       IF #Clr AND NOT #edge THEN
           IF #Q0 THEN #Q0 := FALSE;
           ELSIF #Q1 THEN #Q1 := FALSE;
           ELSIF #Q2 THEN #Q2 := FALSE;
           ELSIF #Q3 THEN #Q3 := FALSE;
           ELSIF #Q4 THEN #Q4 := FALSE;
           ELSIF #Q5 THEN #Q5 := FALSE;
           ELSIF #Q6 THEN #Q6 := FALSE;
           ELSE #Q7 := FALSE;
           END_IF;
       END_IF;
       #edge := #Clr;
   END_IF;


   (* revision history
   hm  25.12.2007  rev 1.0
       original version

   hm  30. oct. 2008   rev 1.1
       optimized performance

   hm  14. mar. 2009   rev 1.2
       removed double assignments

   *)
END_FUNCTION_BLOCK

// ===== PLC "Logic Others"  Unspecific CPU S7 300 =====

FUNCTION_BLOCK "CRC_GEN"   // FB72, SCL
TITLE = CRC_GEN
{ S7_Optimized_Access := 'FALSE' }
AUTHOR : hugo
FAMILY : LOGIC
NAME : CRCGEN
VERSION : 2.0
// CRC_GEN generates a CRC checksum from a block of data and returns  the checksum in a DWORD to be connected to the data for transmission.
// the CRC Polynom is specified with the config variable PN and the length of the Polynom is specified by PL
// A Polynom x4 + X + 1 is represented by 0011 with length 4, the highest order bit is not specified at all..
// The input data is an array of byte of any size, the function is called by CRC_GEN(ADR(array),SIZEOF(array), ....).
// 
// uses: REVERSE (FC310)
//       REFLECT (FC426)
   VAR_INPUT
      PT : Pointer;
      _PT AT PT : Struct
         DBNr : Word;
         Adr : DWord;
      END_STRUCT;
      SIZE : Int;
      PL : Int;
      PN : DWord;
      INIT : DWord;
      REV_IN : Bool;
      REV_OUT : Bool;
      XOR_OUT : DWord;
   END_VAR
   VAR_OUTPUT
      CRC_GEN : DWord;
      _CRC_GEN AT CRC_GEN : Array[0..31] of Bool;
   END_VAR
   VAR_TEMP
      pos : Int;
      shift : Int;
      dx : Byte;
      _dx AT dx : Array[0..7] of Bool;
      bits : Int;
      rTEST_DB : Int;
      Adr : Int;
      DB_LENGTH : Word;
      WRITE_PROT : Bool;
   END_VAR
BEGIN


   (* Datenbaustein Testen *)
   #rTEST_DB := TEST_DB(DB_NUMBER := #_PT.DBNr // IN: WORD
                    ,DB_LENGTH => #DB_LENGTH // OUT: WORD
                    ,WRITE_PROT => #WRITE_PROT // OUT: BOOL
                    ); // INT
   (* Ende wenn Test-DB <> 0 = Fehler *)
   IF #rTEST_DB <> 0 THEN RETURN; END_IF;
   (* Ende wenn DB zu klein *) 
   IF WORD_TO_INT(#DB_LENGTH)/1 < #SIZE THEN RETURN; END_IF;

   #Adr := DWORD_TO_INT(SHR(IN:=SHL(IN:=#_PT.Adr,N:=8),N:=11));

   (* align polygon *)
   #shift := 32 - #PL;
   #PN := SHL(IN:=#PN,N:=#shift);

   (* load first 4 bytes into register minimum message size is 4 bytes
     for smaller messages fill with 0#s at the beginning*)
   FOR #pos := 0 TO 3 DO
     IF #REV_IN THEN #CRC_GEN := SHL(IN:=#CRC_GEN,N:=8) OR "REVERSE"(WORD_TO_BLOCK_DB(#_PT.DBNr).DB(#Adr+#pos)); ELSE #CRC_GEN := SHL(IN:=#CRC_GEN,N:=8) OR WORD_TO_BLOCK_DB(#_PT.DBNr).DB(#Adr+#pos); END_IF;
   END_FOR;
   #pos := 4;

   (* xor with init value *)
   #CRC_GEN := #CRC_GEN XOR SHL(IN:=#INIT,N:=#shift);

   (* calculate CRC for each byte *)
   WHILE #pos < #SIZE DO
     IF #REV_IN THEN #dx := "REVERSE"(WORD_TO_BLOCK_DB(#_PT.DBNr).DB(#Adr+#pos)); ELSE #dx := WORD_TO_BLOCK_DB(#_PT.DBNr).DB(#Adr+#pos); END_IF;
     #pos := #pos + 1;
     (* crc calculation for one byte *)
     FOR #bits := 0 TO 7 DO
       IF #_CRC_GEN[7] THEN
         #CRC_GEN := (SHL(IN:=#CRC_GEN,N:=1) OR BOOL_TO_DWORD(#_dx[7])) XOR #PN;
       ELSE
         #CRC_GEN := SHL(IN:=#CRC_GEN,N:=1) OR BOOL_TO_DWORD(#_dx[7]);
       END_IF;
       #dx := SHL(IN:=#dx,N:=1);
     END_FOR;
   END_WHILE;

   (* all bytes are processed, need to finish the registers 32 bits *)
   FOR #bits := 0 TO 31 DO
     IF #_CRC_GEN[7] THEN
       #CRC_GEN := (SHL(IN:=#CRC_GEN,N:=1) OR BOOL_TO_DWORD(#_dx[7])) XOR #PN;
     ELSE
       #CRC_GEN := SHL(IN:=#CRC_GEN,N:=1) OR BOOL_TO_DWORD(#_dx[7]);
     END_IF;
   END_FOR;

   (* final XOR *)
   #CRC_GEN := SHR(IN:=#CRC_GEN,N:=#shift) XOR #XOR_OUT;

   (* reverse the crc_out put if necessary *)
   IF #REV_OUT THEN #CRC_GEN := "REFLECT"(D:=#CRC_GEN,L:=#PL); END_IF;


   (* typical crc polynoms

   CRC-4-ITU       x4 + x + 1          (ITU G.704, p. 12)  0x3 or 0xC (0x9)
   CRC-5-ITU       x5 + x4 + x2 + 1      (ITU G.704, p. 9)   0x15 or 0x15 (0x0B) Bluetooth
   CRC-5-USB       x5 + x2 + 1         (use: USB token packets)  0x05 or 0x14 (0x9)
   CRC-6-ITU       x6 + x + 1          (ITU G.704, p. 3)   0x03 or 0x30 (0x21)
   CRC-7         x7 + x3 + 1         (use: telecom systems, MMC)   0x09 or 0x48 (0x11)
   CRC-8-ATM       x8 + x2 + x + 1         (use: ATM HEC)  0x07 or 0xE0 (0xC1)
   CRC-8-CCITT     x8 + x7 + x3 + x2 + 1     (use: 1-Wire bus)   0x8D or 0xB1 (0x63)
   CRC-8-Dallas/Maxim  x8 + x5 + x4 + 1      (use: 1-Wire bus)   0x31 or 0x8C (0x19)
   CRC-8         x8 + x7 + x6 + x4 + x2 + 1  0xD5 or 0xAB (0x57)
   CRC-8-SAE J1850   x8 + x4 + x3 + x2 + 1     0x1D or 0xB8
   CRC-10        x10 + x9 + x5 + x4 + x + 1  0x233 or 0x331 (0x263)
   CRC-12        x12 + x11 + x3 + x2 + x + 1 (use: telecom systems)   0x80F or 0xF01 (0xE03)
   CRC-15-CAN      x15 + x14 + x10 + x8 + x7 + x4 + x3 + 1   0x4599 or 0x4CD1 (0x19A3)
   CRC-16-Fletcher   Not a CRC; see Fletcher's checksum  Used in Adler-32 A & B CRCs
   CRC-16-CCITT  x16 + x12 + x5 + 1 (XMODEM,X.25, V.41, Bluetooth, PPP, IrDA; known as "CRC-CCITT")  0x1021 or 0x8408 (0x0811)
   CRC-16-IBM  x16 + x15 + x2 + 1 (USB, many others; also known as "CRC-16")   0x8005 or 0xA001 (0x4003)
   CRC-24-Radix-64   x24 + x23 + x18 + x17 + x14 + x11 + x10 + x7 + x6 + x5 + x4 + x3 + x + 1  0x864CFB or 0xDF3261 (0xBE64C3)
   CRC-32-Adler  Not a CRC; see Adler-32   See Adler-32
   CRC-32-MPEG2  x32 + x26 + x23 + x22 + x16 + x12 + x11 + x10 + x8 + x7 + x5 + x4 + x2 + x + 1  0x04C11DB7 or 0xEDB88320 (0xDB710641) Also used in IEEE 802.3
   CRC-32-IEEE 802.3   x32 + x26 + x23 + x22 + x16 + x12 + x11 + x10 + x8 + x7 + x5 + x4 + x2 + x + 1 (V.42)   0x04C11DB7 or 0xEDB88320 (0xDB710641)
   CRC-32C (Castagnoli)  x32 + x28 + x27 + x26 + x25 + x23 + x22 + x20 + x19 + x18 + x14 + x13 + x11 + x10 + x9 + x8 + x6 + 1  0x1EDC6F41 or 0x82F63B78 (0x05EC76F1)
   CRC-64-ISO  x64 + x4 + x3 + x + 1 (use: ISO 3309)   0x000000000000001B or 0xD800000000000000 (0xB000000000000001)
   CRC-64-ECMA-182   x64 + x62 + x57 + x55 + x54 + x53 + x52 + x47 + x46 + x45 + x40 + x39 + x38 + x37 + x35 + x33 + x32 + x31 + x29 + x27 + x24 + x23 + x22 + x21 + x19 + x17 + x13 + x12 + x10 + x9 + x7 + x4 + x + 1
   (as described in ECMA-182 p.63)   0x42F0E1EBA9EA3693 or 0xC96C5795D7870F42 (0x92D8AF2BAF0E1E85)
   *)



   (* revision history

   hm  9.6.2007    rev 1.0   
     original version 

   hm  11.9.2007   rev 1.1
     deleted unused variable i

   hm  9. oct 2007   rev 1.2
     added init code for crc and xor_out
     added refelct in and reflect_out (rev_in und Rev_out)

   hm  2. jan 2008 rev 1.3
     small changes for performance improvements

   hm  16. mar. 2008 rev 1.4
     changed type of input size to uint

   hm  10. mar. 2009 rev 1.5
     removed nested comments

   hm  16. jan. 2011 rev 2.0
     new version
   *)
END_FUNCTION_BLOCK

FUNCTION_BLOCK "MATRIX"   // FB76, SCL
TITLE = MATRIX
{ S7_Optimized_Access := 'FALSE' }
AUTHOR : hugo
FAMILY : LOGIC
NAME : MATRIX
VERSION : 1.3
// MATRIX is a matrix keyboard encoder for 4 rows and up to 5 columns.
// matrix can send a code while a key is pressed and it sends another code while a key is released when the setup variable 'release' is set to true.
// the setup variable release is false the code is only sent when the key is pressed.
// the output byte holds the 5 columns in the lowest bits 0..2  and the row number in bits 4..6, while bit 7 is true for a key pressed and false for a key released.
   VAR_INPUT
      x1 : Bool;
      x2 : Bool;
      x3 : Bool;
      x4 : Bool;
      X5 : Bool;
      Release : Bool;
   END_VAR
   VAR_OUTPUT
      code : Byte;
      _code AT code : Array[0..7] of Bool;
      TP : Bool;
      y1 : Bool := TRUE;
      y2 : Bool;
      y3 : Bool;
      y4 : Bool;
   END_VAR
   VAR
      line : Byte;
      _line AT line : Array[0..7] of Bool;
      X : Array[0..3] of Byte;
      L : Array[0..3] of Byte;
      i : Int;
      temp : Byte;
      _temp AT temp : Array[0..7] of Bool;
      tempX : Byte;
      _tempX AT tempX : Array[0..7] of Bool;
      tempL : Byte;
      _tempL AT tempL : Array[0..7] of Bool;
   END_VAR
BEGIN


   #TP := FALSE;
   #code := 0;

   (* read scan lines *)
   #tempX := #X[BYTE_TO_INT(#line)];
   #_tempX[0] := #x1;
   #_tempX[1] := #x2;
   #_tempX[2] := #x3;
   #_tempX[3] := #x4;
   #_tempX[4] := #X5;
   #X[BYTE_TO_INT(#line)] := #tempX;

   (* compare for change *)
   FOR #i := 0 TO 3 DO
       IF #X[#i] <> #L[#i] THEN
           (* scan line information has changed code need to be found and generated *)
           #temp := #X[#i] XOR #L[#i];
           #tempX := #X[#i];
           #tempL := #L[#i];
           IF #_temp[0] THEN
               #code := 1;
               #_code[7] := #_tempX[0];
               #_tempL[0] := #_tempX[0];
           ELSIF #_temp[1] THEN
               #code := 2;
               #_code[7] := #_tempX[1];
               #_tempL[1] := #_tempX[1];
           ELSIF #_temp[2] THEN
               #code := 3;
               #_code[7] := #_tempX[2];
               #_tempL[2] := #_tempX[2];
           ELSIF #_temp[3] THEN
               #code := 4;
               #_code[7] := #_tempX[3];
               #_tempL[3] := #_tempX[3];
           ELSIF #_temp[4] THEN
               #code := 5;
               #_code[7] := #_tempX[4];
               #_tempL[4] := #_tempX[4];
           END_IF;
           #X[#i] := #tempX;
           #L[#i] := #tempL;
           #TP := TRUE;
           #_code[4] := #_line[0];
           #_code[5] := #_line[1];
           #_code[6] := #_line[2];

           (* check if release codes need to be killed *)
           IF NOT #Release AND BYTE_TO_INT(#code) < 127 THEN
               #code := 0;
               #TP := FALSE;
           END_IF;
           EXIT;
       END_IF;
   END_FOR;

   (* increment scan line every cycle *)
   #line := INT_TO_BYTE((BYTE_TO_INT(#line) + 1)) AND 2#0000_0011;
   #temp := SHL(IN:=BYTE#1,N:=BYTE_TO_INT(#line));
   #y1 := #_temp[0];
   #y2 := #_temp[1];
   #y3 := #_temp[2];
   #y4 := #_temp[3];




   (* revision history
   hm      10.6.2007   rev 1.0     
       original version 


   hm      11.9.2007   rev 1.1     
       deleted unused variables k and old_code

   hm      23.12.2007  rev 1.2
       added exit statement in for loop instead of i:=5

   hm      26. oct. 2008   rev 1.3
       code optimized

   *)
END_FUNCTION_BLOCK

FUNCTION_BLOCK "PIN_CODE"   // FB233, SCL
TITLE = PIN_CODE
{ S7_Optimized_Access := 'FALSE' }
AUTHOR : hugo
FAMILY : LOOTHER
NAME : PINCODE
VERSION : 1.0
// MATRIX_CODE scans the input of a key_pad (MATRIX) for a sequence of characters.
// 
// uses: CODE [FC229]
//       LEN [FC21]
   VAR_INPUT
      CB : Byte;
      "E" : Bool;
      PIN : String[8];
   END_VAR
   VAR_OUTPUT
      TP : Bool;
   END_VAR
   VAR
      POS : Int := 1;
      CP : Byte;
   END_VAR
BEGIN


   #TP := FALSE;
   IF #"E" THEN
       IF #CB = "CODE"(STR:=#PIN,POS:=#POS) THEN
           #POS := #POS + 1;
           IF #POS > LEN(#PIN) THEN
               (* proper code is detected *)
               #TP := TRUE;
               #POS := 1;
           END_IF;
       ELSE
           #POS := 1;
       END_IF;
   END_IF;


   (* revision history
   hm  30. oct. 2008   rev 1.0     
       original version 


   *)
END_FUNCTION_BLOCK

FUNCTION "CODE" : Byte   // FC229, SCL
TITLE = CODE
{ S7_Optimized_Access := 'FALSE' }
AUTHOR : hugo
FAMILY : STRINGS
NAME : CODE
VERSION : 1.1
// code extracts the code of a character at position POS of a string STR.
   VAR_INPUT
      STR : String[254];
      _STR AT STR : Struct
         length : Byte;
         act_length : Byte;
         str : Array[1..254] of Byte;
      END_STRUCT;
      POS : Int;
   END_VAR
   VAR_TEMP
      PT : Int;   // PT : POINTER TO BYTE;
   END_VAR
BEGIN


   IF #POS < 1 OR #POS > BYTE_TO_INT(#_STR.act_length) THEN
       #CODE := 0;
       RETURN;
   ELSE
       #PT := 1 + (#POS - 1);
       #CODE := #_STR.str[#PT];
   END_IF;

   (* revision history
   hm  9. mar. 2008    rev 1.0
       original version

   hm  29. mar. 2008   rev 1.1
       changed STRING to STRING(STRING_LENGTH)
   *)
END_FUNCTION

FUNCTION "REVERSE" : Byte   // FC310, SCL
TITLE = REVERSE
{ S7_Optimized_Access := 'FALSE' }
AUTHOR : hugo
FAMILY : GATE
NAME : REVERSE
VERSION : 1.1
// This function reverses the bits of a byte so that afdter execution bit 7 is at bit 0 location and so forth.
   VAR_INPUT
      IN : Byte;
   END_VAR
BEGIN


   #REVERSE := SHL(IN:=#IN,N:=7) OR SHR(IN:=#IN,N:=7) OR (ROR(IN:=#IN,N:=3) AND 2#01000100) OR (ROL(IN:=#IN,N:=3) AND 2#00100010)
     OR (SHL(IN:=#IN,N:=1) AND 2#00010000) OR (SHR(IN:=#IN,N:=1) AND 2#00001000);

   (* revision history
   hm    9.oct 2007    rev 1.0
     original version

   hm    18. feb 2008  rev 1.1
     improved performance
   *)
END_FUNCTION

FUNCTION "REFLECT" : DWord   // FC426, SCL
TITLE = REFLECT
{ S7_Optimized_Access := 'FALSE' }
AUTHOR : hugo
FAMILY : GATE
NAME : REFLECT
VERSION : 1.0
// This function reverses the specified amount of bits from bit 0 to bit n within a dword while L specifies the amount of Bits to be reflected.
   VAR_INPUT
      D : DWord;
      L : Int;
   END_VAR
   VAR_TEMP
      tD : DWord;
      i : Int;
   END_VAR
BEGIN


   #tD := #D;
   #REFLECT := 0;
   FOR #i := 1 TO #L DO
     #REFLECT := SHL(IN:=#REFLECT,N:=1) OR (#tD AND DW#16#0000_0001);  //BOOL_TO_DWORD(D.0);
     #tD := SHR(IN:=#tD,N:=1);
   END_FOR;
   #REFLECT := #REFLECT OR SHL(IN:=#tD,N:=#L);


   (* revision history
   hm   16. jan 2011
     new module

   *)
END_FUNCTION

// ===== PLC "Logic gate logic"  Unspecific CPU S7 300 =====

VAR_GLOBAL CONSTANT   // PLC tag table "STEP7 classic symbols"
   "dat" : Byte := 16#1;
   "dat_FC295" : DWord := 16#1;   // MigChange: dat
   "dat_FC297" : Word := 16#1;   // MigChange: dat
END_VAR

FUNCTION_BLOCK "BYTE_TO_BITS"   // FB70, SCL
TITLE = BYTE_TO_BITS
{ S7_Optimized_Access := 'FALSE' }
AUTHOR : hugo
FAMILY : GATE
NAME : BYTE2BIT
VERSION : 1.1
// this Function Block extracts the 8 Bits from a byte
   VAR_INPUT
      IN : Byte;
      tIN AT IN : Array[0..7] of Bool;
   END_VAR
   VAR_OUTPUT
      B0 : Bool;
      B1 : Bool;
      B2 : Bool;
      B3 : Bool;
      B4 : Bool;
      B5 : Bool;
      B6 : Bool;
      B7 : Bool;
   END_VAR
BEGIN


   #B0 := #tIN[0];
   #B1 := #tIN[1];
   #B2 := #tIN[2];
   #B3 := #tIN[3];
   #B4 := #tIN[4];
   #B5 := #tIN[5];
   #B6 := #tIN[6];
   #B7 := #tIN[7];

   (* revision history
   hm    4. aug 2006 rev 1.0
     original version

   hm    16. mar 2008  rev 1.1
     renamed from byte_to_bit to byte_to_bts for compatibility reasons

   *)
END_FUNCTION_BLOCK

FUNCTION_BLOCK "DEC_2"   // FB73, SCL
TITLE = DEC_2
{ S7_Optimized_Access := 'FALSE' }
AUTHOR : hugo
FAMILY : GATE
NAME : DEC_2
VERSION : 1.1
// a bit input will be decoded to the two outputs Q0 or Q1
// dependent on the value of A
// A=0 decodes to Q0 and A=1 decodes to Q1
   VAR_INPUT
      D : Bool;
      "A" : Bool;
   END_VAR
   VAR_OUTPUT
      Q0 : Bool;
      Q1 : Bool;
   END_VAR
BEGIN


     #Q0 := #D AND NOT #"A";
     #Q1 := #D AND #"A";

   (* revision history
   hm 3.3.2007    rev 1.0
       rewritten in ST for better compatibility

   *)
END_FUNCTION_BLOCK

FUNCTION_BLOCK "DEC_4"   // FB74, SCL
TITLE = DEC_4
{ S7_Optimized_Access := 'FALSE' }
AUTHOR : hugo
FAMILY : GATE
NAME : DEC_4
VERSION : 1.1
// a bit input will be decoded to one of the 4 outputs
// dependent on the Adress on A0 and A1
   VAR_INPUT
      D : Bool;
      A0 : Bool;
      A1 : Bool;
   END_VAR
   VAR_OUTPUT
      Q0 : Bool;
      Q1 : Bool;
      Q2 : Bool;
      Q3 : Bool;
   END_VAR
BEGIN


     #Q0 := #D AND NOT #A0 AND NOT #A1;
     #Q1 := #D AND #A0 AND NOT #A1;
     #Q2 := #D AND NOT #A0 AND #A1;
     #Q3 := #D AND #A0 AND #A1;

   (* revision history
   hm 3.3.2007    rev 1.0
       rewritten in ST for better compatibility

   *)
END_FUNCTION_BLOCK

FUNCTION_BLOCK "DEC_8"   // FB75, SCL
TITLE = DEC_8
{ S7_Optimized_Access := 'FALSE' }
AUTHOR : hugo
FAMILY : GATE
NAME : DEC_8
VERSION : 1.3
// a bit input will be decoded to one of the 8 outputs
// dependent on the Adress on A0, A1 and A2
   VAR_INPUT
      D : Bool;
      A0 : Bool;
      A1 : Bool;
      A2 : Bool;
   END_VAR
   VAR_OUTPUT
      Q0 : Bool;
      Q1 : Bool;
      Q2 : Bool;
      Q3 : Bool;
      Q4 : Bool;
      Q5 : Bool;
      Q6 : Bool;
      Q7 : Bool;
   END_VAR
   VAR
      X : Int;
      _X AT X : Array[0..15] of Bool;
   END_VAR
BEGIN


   #X := 0; #_X[8] := #A0; #_X[9] := #A1; #_X[10] := #A2;

   #Q0 := FALSE;
   #Q1 := FALSE; 
   #Q2 := FALSE; 
   #Q3 := FALSE; 
   #Q4 := FALSE; 
   #Q5 := FALSE; 
   #Q6 := FALSE; 
   #Q7 := FALSE;

   CASE #X OF
       0 : #Q0 := #D; 
       1 : #Q1 := #D; 
       2 : #Q2 := #D; 
       3 : #Q3 := #D; 
       4 : #Q4 := #D; 
       5 : #Q5 := #D; 
       6 : #Q6 := #D; 
       7 : #Q7 := #D; 
   END_CASE;


   (* revision history
   hm 3. mar. 2007 rev 1.1
       rewritten in ST for better compatibility

   hm  26. oct. 2008   rev 1.2
       code optimized

   hm  28. mar. 2009   rev 1.3
       replaced multiple assignments
   *)
END_FUNCTION_BLOCK

FUNCTION "BCDC_TO_INT" : Int   // FC290, SCL
TITLE = BCDC_TO_INT
{ S7_Optimized_Access := 'FALSE' }
AUTHOR : hugo
FAMILY : GATE
NAME : BCD2INT
VERSION : 1.1
// this function converts a two digit bcd number into an integer.
   VAR_INPUT
      in : Byte;
   END_VAR
BEGIN


   #BCDC_TO_INT := (BYTE_TO_INT(#in AND 16#0F)) + (WORD_TO_INT(SHR(IN:=BYTE_TO_WORD(#in),N:=4)) * 10);

   (* revision history
   hm  13.12.2007  rev 1.0
       original version

   hm  30.6.2008   rev 1.1
       changed name BCD_TO_INT to BCDC_TO_INT to avoid collision with util.lib

   *)
END_FUNCTION

FUNCTION "BIT_COUNT" : Int   // FC291, SCL
TITLE = BIT_COUNT
{ S7_Optimized_Access := 'FALSE' }
AUTHOR : hugo
FAMILY : GATE
NAME : BITCT
VERSION : 1.1
// BIT_COUNT counts the amount True of bits in a dword.
// for exabple: bit_count(3) returns 2 because two bits (bits 0 and 1) are true and all others are false.
   VAR_INPUT
      IN : DWord;
   END_VAR
   VAR_TEMP
      temp : DWord;
      attemp AT temp : Array[0..31] of Bool;
   END_VAR
BEGIN


     #BIT_COUNT := 0;
     #temp := #IN;

     WHILE DWORD_TO_DINT(#temp) <> 0 DO
       IF #attemp[24] THEN #BIT_COUNT := #BIT_COUNT +1; END_IF;
       #temp := SHR(IN:=#temp,N:=1);
     END_WHILE;

   (* revision history
   5.7.2007  rev 1.0    original version

   10.9.2007  rev 1.1    hm
     changed algorithm for better performace
     the execution time has reduced by a factor of 5
     deleted unused variable temp
   *)
END_FUNCTION

FUNCTION "BIT_LOAD_B" : Byte   // FC292, SCL
TITLE = BIT_LOAD_B
{ S7_Optimized_Access := 'FALSE' }
AUTHOR : hugo
FAMILY : GATE
NAME : BLOADB
VERSION : 1.1
// this function loads a bit into a byte at position pos.
   VAR_INPUT
      IN : Byte;
      VAL : Bool;
      POS : Int;
   END_VAR
BEGIN


   IF #VAL THEN
       #BIT_LOAD_B := #IN OR SHL(IN:="dat",N:=#POS);
   ELSE
       #BIT_LOAD_B := #IN AND (NOT SHL(IN:="dat",N:=#POS));
   END_IF;


   (* revision history
   hm  29. feb 2008    rev 1.0
       original version

   hm  16. mar 2008    rev 1.1
       change input bit to val for compatibility reasons
   *)
END_FUNCTION

FUNCTION "BIT_LOAD_B2" : Byte   // FC294, SCL
TITLE = BIT_LOAD_B2
{ S7_Optimized_Access := 'FALSE' }
AUTHOR : hugo
FAMILY : GATE
NAME : BLOADB2
VERSION : 1.0
// this function loads N bits of D at pos P in Byte I
   VAR_INPUT
      I : Byte;
      D : Bool;
      P : Int;
      N : Int;
   END_VAR
BEGIN


   IF #D THEN
       #BIT_LOAD_B2 := ROL(IN:=SHR(IN:=BYTE#255, N:=8 - #N) OR ROR(IN:=#I, N:=#P), N:=#P);
   ELSE
       #BIT_LOAD_B2 := ROL(IN:=SHL(IN:=BYTE#255, N:=#N) AND ROR(IN:=#I, N:=#P), N:=#P);
   END_IF;



   (* revision history
   hm  18. oct. 2008   rev 1.0
       original version


   *)
END_FUNCTION

FUNCTION "BIT_LOAD_DW" : DWord   // FC295, SCL
TITLE = BIT_LOAD_DW
{ S7_Optimized_Access := 'FALSE' }
AUTHOR : hugo
FAMILY : GATE
NAME : BLOADDW
VERSION : 1.1
// this function loads a bit into a DWord at position pos.
   VAR_INPUT
      IN : DWord;
      VAL : Bool;
      POS : Int;
   END_VAR
BEGIN


   IF #VAL THEN
       #BIT_LOAD_DW := #IN OR SHL(IN:="dat_FC295",N:=#POS);
   ELSE
       #BIT_LOAD_DW := #IN AND (NOT SHL(IN:="dat_FC295",N:=#POS));
   END_IF;


   (* revision history
   hm  29. feb 2008    rev 1.0
       original version

   hm  16. mar 2008    rev 1.1
       change input bit to val for compatibility reasons
   *)
END_FUNCTION

FUNCTION "BIT_LOAD_DW2" : DWord   // FC296, SCL
TITLE = BIT_LOAD_DW2
{ S7_Optimized_Access := 'FALSE' }
AUTHOR : hugo
FAMILY : GATE
NAME : BLOADDW2
VERSION : 1.0
// this function loads N bits of D at pos P in DWORD I
   VAR_INPUT
      I : DWord;
      D : Bool;
      P : Int;
      N : Int;
   END_VAR
BEGIN


   IF #D THEN
       #BIT_LOAD_DW2 := ROL(IN:=SHR(IN:=DWORD#4294967295, N:=32 - #N) OR ROR(IN:=#I, N:=#P), N:=#P);
   ELSE
       #BIT_LOAD_DW2 := ROL(IN:=SHL(IN:=DWORD#4294967295, N:=#N) AND ROR(IN:=#I, N:=#P), N:=#P);
   END_IF;



   (* revision history
   hm  18. oct. 2008   rev 1.0
       original version


   *)
END_FUNCTION

FUNCTION "BIT_LOAD_W" : Word   // FC297, SCL
TITLE = BIT_LOAD_W
{ S7_Optimized_Access := 'FALSE' }
AUTHOR : hugo
FAMILY : GATE
NAME : BLOADW
VERSION : 1.1
// this function loads a bit into a word at position pos.
   VAR_INPUT
      IN : Word;
      VAL : Bool;
      POS : Int;
   END_VAR
BEGIN


   IF #VAL THEN
       #BIT_LOAD_W := #IN OR SHL(IN:="dat_FC297",N:=#POS);
   ELSE
       #BIT_LOAD_W := #IN AND (NOT SHL(IN:="dat_FC297",N:=#POS));
   END_IF;


   (* revision history
   hm  29. feb 2008    rev 1.0
       original version

   hm  16. mar 2008    rev 1.1
       change input bit to val for compatibility reasons
   *)
END_FUNCTION

FUNCTION "BIT_LOAD_W2" : Word   // FC298, SCL
TITLE = BIT_LOAD_W2
{ S7_Optimized_Access := 'FALSE' }
AUTHOR : hugo
FAMILY : GATE
NAME : BLOADW2
VERSION : 1.0
// this function loads N bits of D at pos P in WORD I
   VAR_INPUT
      I : Word;
      D : Bool;
      P : Int;
      N : Int;
   END_VAR
BEGIN


   IF #D THEN
       #BIT_LOAD_W2 := ROL(IN:=SHR(IN:=WORD#65535, N:=16 - #N) OR ROR(IN:=#I, N:=#P), N:=#P);
   ELSE
       #BIT_LOAD_W2 := ROL(IN:=SHL(IN:=WORD#65535, N:=#N) AND ROR(IN:=#I, N:=#P), N:=#P);
   END_IF;



   (* revision history
   hm  18. oct. 2008   rev 1.0
       original version


   *)
END_FUNCTION

FUNCTION "BIT_OF_DWORD" : Bool   // FC299, SCL
TITLE = BIT_OF_DWORD
{ S7_Optimized_Access := 'FALSE' }
AUTHOR : hugo
FAMILY : GATE
NAME : BIToDW
VERSION : 1.2
// this function extracts a single bit from the nth position from right (right is lowest bit)
// the lowest Bit (Bit0 from in) is selected with N=0.
   VAR_INPUT
      IN : DWord;
      N : Int;
   END_VAR
BEGIN


   #BIT_OF_DWORD := DWORD_TO_DINT((SHR(IN:=#IN,N:=#N) AND 16#00000001)) > 0;


   (* old code used before rev 1.1
   temp := SHR(in,n);
   Bit_of_Dword := temp.0;
   *)


   (* revision history
   hm  4. aug. 2006    rev 1.0
       original version

   hm  29. feb 2008    rev 1.1
       improved performance

   hm  6. jun. 2008    rev 1.2
       changes type of input N from byte to int
   *)
END_FUNCTION

FUNCTION "BYTE_OF_BIT" : Byte   // FC300, SCL
TITLE = BYTE_OF_BIT
{ S7_Optimized_Access := 'FALSE' }
AUTHOR : hugo
FAMILY : GATE
NAME : BYTEoBIT
VERSION : 1.1
// this function creates a byte from 8 individual bits
   VAR_INPUT
      B0 : Bool;
      B1 : Bool;
      B2 : Bool;
      B3 : Bool;
      B4 : Bool;
      B5 : Bool;
      B6 : Bool;
      B7 : Bool;
   END_VAR
   VAR_TEMP
      Bx : Byte;
      tBx AT Bx : Array[0..7] of Bool;
   END_VAR
BEGIN


     #tBx[0] := #B0;
     #tBx[1] := #B1;
     #tBx[2] := #B2;
     #tBx[3] := #B3;
     #tBx[4] := #B4;
     #tBx[5] := #B5;
     #tBx[6] := #B6;
     #tBx[7] := #B7;

     #BYTE_OF_BIT := #Bx;

   (* original code
   Byte_of_bit := SHL(SHL(SHL(SHL(SHL(SHL(SHL(BOOL_TO_BYTE(B7),1) OR BOOL_TO_BYTE(B6),1) OR BOOL_TO_BYTE(B5),1) OR BOOL_TO_BYTE(B4),1)
     OR BOOL_TO_BYTE(B3),1) OR BOOL_TO_BYTE(B2),1) OR BOOL_TO_BYTE(B1),1) OR BOOL_TO_BYTE(B0);
   *)

   (* revision history

   hm  4. aug 2006   rev 1.0
     original version

   hm  18. feb. 2008 rev 1.1
     improved performance

   *)
END_FUNCTION

FUNCTION "BYTE_OF_DWORD" : Byte   // FC301, SCL
TITLE = BYTE_OF_DWORD
{ S7_Optimized_Access := 'FALSE' }
AUTHOR : hugo
FAMILY : GATE
NAME : BYTEoDW
VERSION : 1.2
// this function extracts a single byte from the nth position from right (right is lowest byte) 
// the lower byte (starting with Bit0 from in) is selected with N=0.
   VAR_INPUT
      in : DWord;
      N : Int;
   END_VAR
BEGIN


   #BYTE_OF_DWORD := DWORD_TO_BYTE(SHR(IN:=#in,N:=WORD_TO_INT(SHL(IN:=INT_TO_WORD(#N),N:=3))));

   (* revision history
   hm  17. jan 2007    rev 1.0
       original version

   hm  2. jan 2008     rev 1.1
       improved performance

   hm  30. oct. 2008   rev 1.2
       improved performance
   *)
END_FUNCTION

FUNCTION "CHECK_PARITY" : Bool   // FC302, SCL
TITLE = CHECK_PARITY
{ S7_Optimized_Access := 'FALSE' }
AUTHOR : hugo
FAMILY : GATE
NAME : CHECKP
VERSION : 1.3
// this function checks for an even partity for a dword and partity bit.
   VAR_INPUT
      in : DWord;
      p : Bool;
   END_VAR
   VAR_TEMP
      cnt : Int;
      tIN : DWord;
      _IN AT tIN : Array[0..31] of Bool;
   END_VAR
BEGIN


     #tIN := #in;
     #cnt := 0;

     #CHECK_PARITY := NOT #p;

     WHILE #tIN <> 0 DO
       #CHECK_PARITY := #CHECK_PARITY XOR #_IN[24] XOR #_IN[25] XOR #_IN[26] XOR #_IN[27];
       #tIN := SHR(IN:=#tIN,N:=4);
     END_WHILE;

   (* code before rev 1.2
   WHILE in > 0 DO
     IF in.0 THEN cnt := cnt + 1; END_IF;
     in := SHR(in,1);
   END_WHILE;
   check_parity := even(cnt) XOR P;
   *)


   (* revision history

   rev 1.0 HM  1.oct.2006

   rev 1.1 hm  10.sep.2007
     changed algorithm to improove performance

   rev 1.2 hm  8 dec 2007
     changed algorithm to improove performance

   rev 1.3 hm  18. feb 2008
     changed algorithm to improove performance
   *)
END_FUNCTION

FUNCTION "DW_TO_REAL" : Real   // FC303, SCL
TITLE = DW_TO_REAL
{ S7_Optimized_Access := 'FALSE' }
AUTHOR : hugo
FAMILY : GATE
NAME : BIT2REAL
VERSION : 1.0
// this function converts a DWORD to REAL in a bitwise manner.
   VAR_INPUT
      X : DWord;
   END_VAR
BEGIN


   //pt := ADR(X);
   #DW_TO_REAL := DWORD_TO_REAL(#X);    //pt^;

   (* revision history
   hm  18. apr. 2008
       original version

   *)
END_FUNCTION

FUNCTION "DWORD_OF_BYTE" : DWord   // FC304, SCL
TITLE = DWORD_OF_BYTE
{ S7_Optimized_Access := 'FALSE' }
AUTHOR : hugo
FAMILY : GATE
NAME : DWoBYTE
VERSION : 1.3
// this function creates a Dword from 4 individual bytes
   VAR_INPUT
      B3 : Byte;
      B2 : Byte;
      B1 : Byte;
      B0 : Byte;
   END_VAR
BEGIN


   #DWORD_OF_BYTE := SHL(IN:=SHL(IN:=SHL(IN:=BYTE_TO_DWORD(#B3),N:=8) OR BYTE_TO_DWORD(#B2),N:=8) OR BYTE_TO_DWORD(#B1),N:=8) OR BYTE_TO_DWORD(#B0);


   (* revision history
   hm  24. jan 2007  rev 1.0
     original version

   hm 2. jan 2008  rev 1.1
     inproved performance

   hm  23. apr. 2008 rev 1.2
     reverse order of inputs to be more logical

   hm  18. jul. 2009 rev 1.3
     added type conversions for compatibility reasons
   *)
END_FUNCTION

FUNCTION "INT_TO_BCDC" : Byte   // FC305, SCL
TITLE = INT_TO_BCDC
{ S7_Optimized_Access := 'FALSE' }
AUTHOR : hugo
FAMILY : GATE
NAME : INT2BCD
VERSION : 1.1
// this function converts an integer into a two digit bcd number.
   VAR_INPUT
      IN : Int;
   END_VAR
BEGIN


   #INT_TO_BCDC := SHL(IN:=INT_TO_BYTE(#IN / INT#10),N:=4) OR INT_TO_BYTE(#IN MOD INT#10);

   (* revision history
   hm  13.12.2007
       original version

   hm  30.6.2008   rev 1.1
       changed name INT_TO_BCD to INT_TO_BCDC to avoid collision with util.lib
       corrected error in code

   *)
END_FUNCTION

FUNCTION "MUX_2" : Bool   // FC306, SCL
TITLE = MUX_2
{ S7_Optimized_Access := 'FALSE' }
AUTHOR : hugo
FAMILY : GATE
NAME : MUX_2
VERSION : 1.2
// dual input multiplexer
// depending on the value of A0, D0 or D1 will be switched to the Output
   VAR_INPUT
      D0 : Bool;
      D1 : Bool;
      A0 : Bool;
   END_VAR
BEGIN


   #MUX_2 := SEL(G:=#A0, IN0:=#D0, IN1:=#D1);


   (*
   revision history:
   hm  5.10.2006       rev 1.1
       changed to ST Langage for better portability.

   hm  16. oct. 2008   rev 1.2
       improved performance

   *)
END_FUNCTION

FUNCTION "MUX_4" : Bool   // FC307, SCL
TITLE = MUX_4
{ S7_Optimized_Access := 'FALSE' }
AUTHOR : hugo
FAMILY : GATE
NAME : MUX_4
VERSION : 1.2
// quad input multiplexer
// depending on the value of A0 and A1, one of the 4 inputs will be switched to the Output
   VAR_INPUT
      D0 : Bool;
      D1 : Bool;
      D2 : Bool;
      D3 : Bool;
      A0 : Bool;
      A1 : Bool;
   END_VAR
BEGIN


   IF #A1 THEN
       #MUX_4 := SEL(G:=#A0, IN0:=#D2, IN1:=#D3);
   ELSE
       #MUX_4 := SEL(G:=#A0, IN0:=#D0, IN1:=#D1);
   END_IF;

   (*
   revision history:
   hm  5.10.2006       rev 1.1
       rewritten to ST for better portability

   hm  16. oct. 2008   rev 1.2
       improved performance

   *)
END_FUNCTION

FUNCTION "PARITY" : Bool   // FC308, SCL
TITLE = PARITY
{ S7_Optimized_Access := 'FALSE' }
AUTHOR : hugo
FAMILY : GATE
NAME : PARITY
VERSION : 1.3
// this function calculates the even parity of an input Dword
// the output will be true if the amount of high bits are an odd number.
   VAR_INPUT
      in : DWord;
   END_VAR
   VAR_TEMP
      tIN : DWord;
      _IN AT tIN : Array[0..31] of Bool;
   END_VAR
BEGIN


     #tIN := #in;
     #PARITY := 0;

     WHILE #tIN <> 0 DO
       #PARITY := #PARITY XOR #_IN[24] XOR #_IN[25] XOR #_IN[26] XOR #_IN[27];
       #tIN := SHR(IN:=#tIN,N:=4);
     END_WHILE;


   (* code before rev 1.2
   WHILE in > 0 DO
     IF in.0 THEN cnt := cnt +1; END_IF;
     in := SHR(in,1);
   END_WHILE;
   IF (cnt MOD 2) = 1 THEN parity := TRUE; ELSE parity := FALSE; END_IF;
   *)

   (* revision history

   rev 1.0 hm 1 sep 2006
     original version

   rev 1.1 hm 10.9.2007
     changed algorithm to improve performance

   rev 1.2 hm  8 dec 2007
     changed algorithm to improve performance

   rev 1.3 hm  18 feb 2008
     changed algorithm to improve performance
   *)
END_FUNCTION

FUNCTION "REAL_TO_DW" : DWord   // FC309, SCL
TITLE = REAL_TO_DW
{ S7_Optimized_Access := 'FALSE' }
AUTHOR : hugo
FAMILY : GATE
NAME : REAL2BIT
VERSION : 1.0
// this function converts a 32 Bit Real to a dword in a bitwise manner.
   VAR_INPUT
      X : Real;
   END_VAR
BEGIN


   //pt := ADR(X);
   #REAL_TO_DW := REAL_TO_DWORD(#X);    //pt^;

   (* revision history
   hm  18. apr. 2008
       original version

   *)
END_FUNCTION

FUNCTION "REVERSE" : Byte   // FC310, SCL
TITLE = REVERSE
{ S7_Optimized_Access := 'FALSE' }
AUTHOR : hugo
FAMILY : GATE
NAME : REVERSE
VERSION : 1.1
// This function reverses the bits of a byte so that afdter execution bit 7 is at bit 0 location and so forth.
   VAR_INPUT
      IN : Byte;
   END_VAR
BEGIN


   #REVERSE := SHL(IN:=#IN,N:=7) OR SHR(IN:=#IN,N:=7) OR (ROR(IN:=#IN,N:=3) AND 2#01000100) OR (ROL(IN:=#IN,N:=3) AND 2#00100010)
     OR (SHL(IN:=#IN,N:=1) AND 2#00010000) OR (SHR(IN:=#IN,N:=1) AND 2#00001000);

   (* revision history
   hm    9.oct 2007    rev 1.0
     original version

   hm    18. feb 2008  rev 1.1
     improved performance
   *)
END_FUNCTION

FUNCTION "SHL1" : DWord   // FC311, SCL
TITLE = SHL1
{ S7_Optimized_Access := 'FALSE' }
AUTHOR : hugo
FAMILY : GATE
NAME : SHL1
VERSION : 1.1
// SHL1 shifts N bits to the left filling the new bits with 1
   VAR_INPUT
      IN : DWord;
      N : Int;
   END_VAR
   VAR_TEMP
      temp : DWord;
   END_VAR
BEGIN


     #temp := 16#FFFF_FFFF;

     #SHL1 := SHR(IN:=#temp,N:=32-#N) OR SHL(IN:=#IN,N:=#N);

   (* revision history
   hm  14.9.2007   rev 1.0
     original version

   hm  27. dec 2007  rev 1.1
     changed code for better performance

   *)
END_FUNCTION

FUNCTION "SHR1" : DWord   // FC312, SCL
TITLE = SHR1
{ S7_Optimized_Access := 'FALSE' }
AUTHOR : hugo
FAMILY : GATE
NAME : SHR1
VERSION : 1.1
// SHR1 shifts N bits to the right filling the new bits with 1
   VAR_INPUT
      IN : DWord;
      N : Int;
   END_VAR
   VAR_TEMP
      temp : DWord;
   END_VAR
BEGIN


     #temp := 16#FFFF_FFFF;

     #SHR1 := SHL(IN:=#temp,N:=32-#N) OR SHR(IN:=#IN,N:=#N);

   (* revision history
   hm  14.9.2007   rev 1.0
     original version

   hm  27. dec 2007  rev 1.1
     changed code for better performance

   *)
END_FUNCTION

FUNCTION "SWAP_BYTE" : Word   // FC313, SCL
TITLE = SWAP_BYTE
{ S7_Optimized_Access := 'FALSE' }
AUTHOR : hugo
FAMILY : GATE
NAME : SWAPBY
VERSION : 1.0
// This function swaps the high and low byte of the word in.
   VAR_INPUT
      IN : Word;
   END_VAR
BEGIN


     #SWAP_BYTE := ROL(IN:=#IN,N:=8);


   (* revision history
   hm    4. feb 2008 rev 1.0
     original version

   *)
END_FUNCTION

FUNCTION "SWAP_BYTE2" : DWord   // FC314, SCL
TITLE = SWAP_BYTE2
{ S7_Optimized_Access := 'FALSE' }
AUTHOR : hugo
FAMILY : GATE
NAME : SWAPBY2
VERSION : 1.0
// This function reverses the byte order in the dword.
   VAR_INPUT
      IN : DWord;
   END_VAR
BEGIN


     #SWAP_BYTE2 := (ROR(IN:=#IN,N:=8) AND 16#FF00FF00) OR (ROL(IN:=#IN,N:=8) AND 16#00FF00FF);

   (* revision history
   hm    4. feb 2008 rev 1.0
     original version

   *)
END_FUNCTION

FUNCTION "WORD_OF_BYTE" : Word   // FC315, SCL
TITLE = WORD_OF_BYTE
{ S7_Optimized_Access := 'FALSE' }
AUTHOR : hugo
FAMILY : GATE
NAME : WoBYTE
VERSION : 1.4
// this function creates a word from 2 individual bytes
   VAR_INPUT
      B1 : Byte;
      B0 : Byte;
   END_VAR
BEGIN


   #WORD_OF_BYTE := SHL(IN:=BYTE_TO_WORD(#B1),N:=8) OR BYTE_TO_WORD(#B0);


   (* revision history
   hm  24. jan 2007  rev 1.0
     original version

   hm  2. jan 2008 rev 1.1
     improved performance

   hm  19. feb 2008  rev 1.2
     replaced and with or for better compatibility

   hm  23. apr. 2008 rev 1.3
     reverse order of inputs to be more logical

   hm  18. jul. 2009 rev 1.4
     added type conversions for compatibility reasons

   *)
END_FUNCTION

FUNCTION "WORD_OF_DWORD" : Word   // FC316, SCL
TITLE = WORD_OF_DWORD
{ S7_Optimized_Access := 'FALSE' }
AUTHOR : hugo
FAMILY : GATE
NAME : WoDW
VERSION : 1.2
// this function extracts a single word from the nth position from right (right is lowest byte)
// the lower word (starting weith Bit0 from in) is selected with N=0.
   VAR_INPUT
      in : DWord;
      N : Int;
   END_VAR
BEGIN


   #WORD_OF_DWORD := DWORD_TO_WORD(SHR(IN:=#in,N:=WORD_TO_INT(SHL(IN:=INT_TO_WORD(#N),N:=4))));

   (* revision history
   hm  17. jan 2007    rev 1.0
       original version

   hm  2. jan 2008     rev 1.1
       improved performance

   hm  30. oct. 2008   rev 1.2
       improved performance
   *)
END_FUNCTION

FUNCTION "BIT_TOGGLE_W" : Word   // FC396, SCL
TITLE = BIT_TOGGLE_W
{ S7_Optimized_Access := 'FALSE' }
AUTHOR : hugo
FAMILY : GATE
NAME : BITTOGW
VERSION : 1.0
// this function toggles a bit of a WORD at position pos.
   VAR_INPUT
      IN : Word;
      POS : Int;
   END_VAR
BEGIN


   #BIT_TOGGLE_W := SHL(IN:=WORD#1, N:=#POS) XOR #IN;



   (* revision history
   hm  18. oct. 2008   rev 1.0
       original version


   *)
END_FUNCTION

FUNCTION "BIT_TOGGLE_B" : Byte   // FC397, SCL
TITLE = BIT_TOGGLE_B
{ S7_Optimized_Access := 'FALSE' }
AUTHOR : hugo
FAMILY : GATE
NAME : BITTOGB
VERSION : 1.0
// this function toggles a bit of a BYTE at position pos.
   VAR_INPUT
      IN : Byte;
      POS : Int;
   END_VAR
BEGIN


   #BIT_TOGGLE_B := SHL(IN:=BYTE#1, N:=#POS) XOR #IN;




   (* revision history
   hm  18. oct. 2008   rev 1.0
       original version


   *)
END_FUNCTION

FUNCTION "BIT_TOGGLE_DW" : DWord   // FC398, SCL
TITLE = BIT_TOGGLE_DW
{ S7_Optimized_Access := 'FALSE' }
AUTHOR : hugo
FAMILY : GATE
NAME : BITTOGDW
VERSION : 1.0
// this function toggles a bit of a WORD at position pos.
   VAR_INPUT
      IN : DWord;
      POS : Int;
   END_VAR
BEGIN


   #BIT_TOGGLE_DW := SHL(IN:=DWORD#1, N:=#POS) XOR #IN;



   (* revision history
   hm  18. oct. 2008   rev 1.0
       original version


   *)
END_FUNCTION

FUNCTION "DWORD_OF_WORD" : DWord   // FC419, SCL
TITLE = DWORD_OF_WORD
{ S7_Optimized_Access := 'FALSE' }
AUTHOR : hugo
FAMILY : GATE
NAME : DWoWORD
VERSION : 1.0
// this function creates a Dword from 2 individual Words
   VAR_INPUT
      W1 : Word;
      W0 : Word;
   END_VAR
BEGIN


   #DWORD_OF_WORD := SHL(IN:=WORD_TO_DWORD(#W1),N:=16) OR WORD_TO_DWORD(#W0);


   (* revision history

   hm  18. jul. 2009 rev 1.0
     original version

   *)
END_FUNCTION

FUNCTION "BYTE_TO_GRAY" : Byte   // FC420, SCL
TITLE = BYTE_TO_GRAY
{ S7_Optimized_Access := 'FALSE' }
AUTHOR : hugo
FAMILY : GATE
NAME : BY2GRAY
VERSION : 1.0
// this function converts a binary to gray code
   VAR_INPUT
      IN : Byte;
   END_VAR
BEGIN


   #BYTE_TO_GRAY := #IN XOR SHR(IN:=#IN,N:=1);

   (* revision history
   hm  9. nov. 2009  rev 1.0
     original version

   *)
END_FUNCTION

FUNCTION "GRAY_TO_BYTE" : Byte   // FC421, SCL
TITLE = GRAY_TO_BYTE
{ S7_Optimized_Access := 'FALSE' }
AUTHOR : hugo
FAMILY : GATE
NAME : GRAY2BY
VERSION : 1.0
// this function converts a gray code into binary
   VAR_INPUT
      IN : Byte;
   END_VAR
BEGIN


   #GRAY_TO_BYTE := SHR(IN:=#IN,N:=4) XOR #IN;
   #GRAY_TO_BYTE := SHR(IN:=#GRAY_TO_BYTE,N:=2) XOR #GRAY_TO_BYTE;
   #GRAY_TO_BYTE := SHR(IN:=#GRAY_TO_BYTE,N:=1) XOR #GRAY_TO_BYTE;

   (* revision history
   hm  9. nov. 2009  rev 1.0
     original version

   *)
END_FUNCTION

FUNCTION "CHK_REAL" : Byte   // FC425, SCL
TITLE = CHK_REAL
{ S7_Optimized_Access := 'FALSE' }
AUTHOR : hugo
FAMILY : GATE
NAME : CHKREAL
VERSION : 1.0
// this function checks a floating point variable of type real (IEEE754-32Bits) for NAN and infinity
// RETURN values: #0 = normal value, #20 = +infinity, #40 = -infinty, #80 = NAN
   VAR_INPUT
      X : Real;
   END_VAR
   VAR_TEMP
      pt : DWord;
      tmp : DWord;
   END_VAR
BEGIN


   #pt := REAL_TO_DWORD(#X);       (* move real to dword, real_to_dword does not work becasze it treats dword as a number on many systems *)
   #tmp := ROL(IN:=#pt,N:=1);      (* rotate left foir easy checking, sign will be at lease significant digit *)
   IF DWORD_TO_DINT(#tmp) < DWORD_TO_DINT(16#FF000000) THEN
     #CHK_REAL := 16#00;    (* normalized and denormalized numbers *)
   ELSIF #tmp = 16#FF000000 THEN
     #CHK_REAL := 16#20;    (* X is +infinity see IEEE754 *)
   ELSIF #tmp = 16#FF000001 THEN
     #CHK_REAL := 16#40;    (* X is -infinity see IEEE754 *)
   ELSE
     #CHK_REAL := 16#80;    (* X is NAN see IEEE754 *)
   END_IF;


   (* revision history
   hm   20. jan. 2011  rev 1.0
     original version

   *)
END_FUNCTION

FUNCTION "REFLECT" : DWord   // FC426, SCL
TITLE = REFLECT
{ S7_Optimized_Access := 'FALSE' }
AUTHOR : hugo
FAMILY : GATE
NAME : REFLECT
VERSION : 1.0
// This function reverses the specified amount of bits from bit 0 to bit n within a dword while L specifies the amount of Bits to be reflected.
   VAR_INPUT
      D : DWord;
      L : Int;
   END_VAR
   VAR_TEMP
      tD : DWord;
      i : Int;
   END_VAR
BEGIN


   #tD := #D;
   #REFLECT := 0;
   FOR #i := 1 TO #L DO
     #REFLECT := SHL(IN:=#REFLECT,N:=1) OR (#tD AND DW#16#0000_0001);  //BOOL_TO_DWORD(D.0);
     #tD := SHR(IN:=#tD,N:=1);
   END_FOR;
   #REFLECT := #REFLECT OR SHL(IN:=#tD,N:=#L);


   (* revision history
   hm   16. jan 2011
     new module

   *)
END_FUNCTION

// ===== PLC "Logic generators"  Unspecific CPU S7 300 =====

VAR_GLOBAL CONSTANT   // PLC tag table "STEP7 classic symbols"
   "debug" : Bool := FALSE;
   "N" : Int := 0;
   "offset" : Int := 0;
   "offset_1" : DWord := 0;
END_VAR

DATA_BLOCK "IDB_STIME"   // DB64
{ S7_Optimized_Access := 'FALSE' }
AUTHOR : dalbi
FAMILY : MEASURE
VERSION : 0.0
// stored: InstanceOfName STIME
"STIME"
BEGIN
END_DATA_BLOCK

FUNCTION_BLOCK "A_TRIG"   // FB41, SCL
TITLE = A_TRIG
{ S7_Optimized_Access := 'FALSE' }
AUTHOR : hugo
FAMILY : GENERAT
NAME : A_TRIG
VERSION : 1.1
// this block is similar to the IEC Standard R_trig and F_trig but it monitors a REAL for change.
// if the valiue on IN changes more then D from the last value it will generate trigger and display the difference in output D.
// the trigger will only be active for one cycle.
   VAR_INPUT
      IN : Real;
      RES : Real;
   END_VAR
   VAR_OUTPUT
      Q : Bool;
      D : Real;
   END_VAR
   VAR
      last_in : Real;
   END_VAR
BEGIN


   #D:= #IN - #last_in;
   #Q := ABS(#D) > #RES;
   IF #Q THEN #last_in := #IN; END_IF;
   #D := #IN - #last_in;


   (* revision history

   hm  16. jul. 2008   rev 1.0
       original version released

   hm  25. oct. 2008   rev 1.1
       code optimization
       a_trig now also works for res = 0

   *)
END_FUNCTION_BLOCK

FUNCTION_BLOCK "B_TRIG"   // FB42, SCL
TITLE = B_TRIG
{ S7_Optimized_Access := 'FALSE' }
AUTHOR : hugo
FAMILY : GENERAT
NAME : B_TRIG
VERSION : 1.0
// this block is similar to R_trig and F_trig but it generates a pulse on rising and falling edge.
   VAR_INPUT
      CLK : Bool;
   END_VAR
   VAR_OUTPUT
      Q : Bool;
   END_VAR
   VAR
      edge : Bool;
   END_VAR
BEGIN


     #Q := #CLK XOR #edge;
     #edge := #CLK;
END_FUNCTION_BLOCK

FUNCTION_BLOCK "CLICK_CNT"   // FB43, SCL
TITLE = CLICK_CNT
{ S7_Optimized_Access := 'FALSE' }
AUTHOR : hugo
FAMILY : GENERAT
NAME : CLICKCNT
VERSION : 1.0
// this Module decodes a specified number of clicks.
// the output trig is high for one cycle if N clicks are present within a specified time TC.
   VAR_INPUT
      IN : Bool;
      N : Int;
      TC : Time;
   END_VAR
   VAR_OUTPUT
      Q : Bool;
   END_VAR
   VAR
      tx : TP;
      edge : Bool;
      cnt : Int := -1;
   END_VAR
BEGIN


   (* Q shall only be active for one cycle only *)
   #Q := FALSE;


   IF #IN AND NOT #edge AND NOT #tx.Q THEN
       (* a rising edge on in sets the counter to 0 *)
       #cnt := 0;
   ELSIF #tx.Q AND NOT #IN AND #edge THEN
       (* count falling edges when tp.q is true *)
       #cnt := #cnt + 1;
   ELSIF NOT #tx.Q THEN
       #Q := #cnt = #N;
       #cnt := -1;
   END_IF;

   (* remember the status of IN *)
   #edge := #IN;
   #tx(IN := #IN, PT := #TC);


   (* revision history

   hm  16. jul. 2008   rev 1.0
       original version released


   *)
END_FUNCTION_BLOCK

FUNCTION_BLOCK "CLICK_DEC"   // FB44, SCL
TITLE = CLICK_DEC
{ S7_Optimized_Access := 'FALSE' }
AUTHOR : hugo
FAMILY : GENERAT
NAME : CLICKDEC
VERSION : 1.1
// this Module detects a rising edge on In and decodes the amount of falling edges (Pulses) within a specified time TC.
// the outputs Q0..Q3 will go true for one cycle and the amount of clicks within a specified time TC.
// if only a rising egde is detected within TC Q0 will respond, Q1 for 1 pulse and so on..
   VAR_INPUT
      IN : Bool;
      TC : Time;
   END_VAR
   VAR_OUTPUT
      Q0 : Bool;
      Q1 : Bool;
      Q2 : Bool;
      Q3 : Bool;
   END_VAR
   VAR
      tx : TP;
      edge : Bool;
      cnt : Int := -1;
   END_VAR
BEGIN


   (* Q shall only be active for one cycle only *)
   IF #IN = FALSE THEN
       #Q3 := FALSE;
       #Q2 := FALSE;
       #Q1 := FALSE;
       #Q0 := FALSE; 
   END_IF;

   IF #IN AND NOT #edge AND NOT #tx.Q THEN
       (* a rising edge on in sets the counter to 0 *)
       #cnt := 0;
   ELSIF #tx.Q AND NOT #IN AND #edge THEN
       (* count falling edges when tp.q is true *)
       #cnt := #cnt + 1;
   ELSIF NOT #tx.Q THEN
       CASE #cnt OF
           0 : #Q0 := TRUE;
           1 : #Q1 := TRUE;
           2 : #Q2 := TRUE;
           3 : #Q3 := TRUE;
       END_CASE;
       #cnt := -1;
   END_IF;

   (* remember the status of IN *)
   #edge := #IN;
   #tx(IN := #IN, PT := #TC);


   (* revision history

   hm 17. jul. 2008    rev 1.0
       original version released

   hm  14. mar. 2009   rev 1.1
       removed double assignments

   *)
END_FUNCTION_BLOCK

FUNCTION_BLOCK "CLK_DIV"   // FB50, SCL
TITLE = CLK_DIV
{ S7_Optimized_Access := 'FALSE' }
AUTHOR : hugo
FAMILY : GENERAT
NAME : CLK_DIV
VERSION : 1.1
// this is a clock divider
// each output divides the signal by 2
// Q0 = clk / 2 , Q1 = Q0 / 2 and so on.
// the outputs have a 50% duty cycle each.
   VAR_INPUT
      clk : Bool;
      rst : Bool;
   END_VAR
   VAR_OUTPUT
      Q0 : Bool;
      Q1 : Bool;
      Q2 : Bool;
      Q3 : Bool;
      Q4 : Bool;
      Q5 : Bool;
      Q6 : Bool;
      Q7 : Bool;
   END_VAR
   VAR
      cnt : Byte;
      _cnt AT cnt : Array[0..7] of Bool;
   END_VAR
BEGIN


   IF #rst THEN
       #cnt:= 0;
       #Q0 := 0;
       #Q1 := 0;
       #Q2 := 0;
       #Q3 := 0;
       #Q4 := 0;
       #Q5 := 0;
       #Q6 := 0;
       #Q7 := 0;
   ELSIF #clk THEN
       #cnt:= INT_TO_BYTE(BYTE_TO_INT(#cnt) +1);
       #Q0 := #_cnt[0];
       #Q1 := #_cnt[1];
       #Q2 := #_cnt[2];
       #Q3 := #_cnt[3];
       #Q4 := #_cnt[4];
       #Q5 := #_cnt[5];
       #Q6 := #_cnt[6];
       #Q7 := #_cnt[7];
   END_IF;


   (* revision history
   hm  4. aug. 2006  rev 1.0
     original version

   hm  2. jan 2008   rev 1.1
     improved performance

   *)
END_FUNCTION_BLOCK

FUNCTION_BLOCK "CLK_N"   // FB51, SCL
TITLE = CLK_N
{ S7_Optimized_Access := 'FALSE' }
AUTHOR : hugo
FAMILY : GENERAT
NAME : CLK_N
VERSION : 1.0
// clk_N uses the internal sps time to generate one pulse every N ms
// every pulse is only valid for one cycle so that a edge trigger is not necessary
// clk_N generates pulses depending on the accuracy of the system clock.
// The input N controlls the period time of the clock.
// N=0 equals 1ms, N=1 equals 2ms, N=2 equals 4ms, N=3 equals 8ms ....
//  
// be careful, 1ms clocks will only work on very powerful sps cpu's
// 
// uses: T_PLC_MS [FC64]
//       STIME [FB64],IDB_STIME [DB64]
   VAR_INPUT
      N : Int;
   END_VAR
   VAR_OUTPUT
      Q : Bool;
   END_VAR
   VAR
      edge : Bool;
      stime : DWord;
      _stime AT stime : Array[0..31] of Bool;
      clk : Bool;
   END_VAR
BEGIN


     #stime := SHR(IN:="T_PLC_MS"(),N:=#N);
     #clk := #_stime[24]; // .0
     #Q := #clk XOR #edge;
     #edge := #clk;

   (* revision history
   hm  16. dec 2007    rev 1.0
     original version

   *)
END_FUNCTION_BLOCK

FUNCTION_BLOCK "CLK_PRG"   // FB52, SCL
TITLE = CLK_PRG
{ S7_Optimized_Access := 'FALSE' }
AUTHOR : hugo
FAMILY : GENERAT
NAME : CLK_PRG
VERSION : 1.3
// clk_prg uses the internal sps time to generate a clock with programmable period time.
// the period time is defined for 10ms .. 65s
// the first cycle after start is a clk pulse and then depending on the programmed period time a delay.
// every pulse is only valid for one cycle.
// the accuracy of clk_prg is depending on the accuracy of the system clock.
// 
// uses: T_PLC_MS [FC64]
//       STIME [FB64],IDB_STIME [DB64]
   VAR_INPUT
      PT : Time := T#10MS;
   END_VAR
   VAR_OUTPUT
      Q : Bool;
   END_VAR
   VAR
      init : Bool;
      last : Time;
      tx : Time;
   END_VAR
   VAR_TEMP
      TOP_SI : Struct
         EV_CLASS : Byte;
         EV_NUM : Byte;
         PRIORITY : Byte;
         NUM : Byte;
         TYP2_3 : Byte;
         TYP1 : Byte;
         ZI1 : Word;
         ZI2_3 : DWord;
      END_STRUCT;
      START_UP_SI : Struct
         EV_CLASS : Byte;
         EV_NUM : Byte;
         PRIORITY : Byte;
         NUM : Byte;
         TYP2_3 : Byte;
         TYP1 : Byte;
         ZI1 : Word;
         ZI2_3 : DWord;
      END_STRUCT;
      ERR : Int;
   END_VAR
BEGIN


   (* read actual startup info *)
   (* OB1_SCAN_1  BYTE  -  B#16#01: Abschluss des Neustarts (Warmstarts)
                        -  B#16#02: Abschluss des Wiederanlaufs
                        -  B#16#03: Abschluss des freien Zyklus
                        -  B#16#04: Abschluss des Kaltstarts
                        -  B#16#05: Erster OB 1-Zyklus der neuen Master-CPU nach 
                                    Master-Reserve-Umschaltung und STOP des 
                                    bisherigen Masters *)

   #ERR := RD_SINFO (TOP_SI => #TOP_SI, START_UP_SI => #START_UP_SI);

   (* read system time *)
   #tx := T_CONV(DWORD_TO_DINT("T_PLC_MS"()));

   (* reset last_time on system startup *)
   IF #TOP_SI.EV_NUM = 1 OR #TOP_SI.EV_NUM = 2 OR #TOP_SI.EV_NUM = 4 THEN 
       #init := false;
   END_IF;

   (* initialize on startup *)
   IF NOT #init THEN
       #init := TRUE;
       #last := #tx - #PT;
   END_IF;

   (* generate output pulse when next_pulse is reached *)
   #Q := #tx - #last >= #PT;
   IF #Q THEN #last := #tx; END_IF;


   (* revision hiostory

   hm 25 feb 2007  rev 1.1
       rewritten code for higher performance
       pt can now be changed during runtime

   hm  17. sep 2007    rev 1.2
       replaced time() with t_plc_ms() for compatibility reasons

   hm  25. oct. 2008   rev 1.3
       optimized code

   *)
END_FUNCTION_BLOCK

FUNCTION_BLOCK "CLK_PULSE"   // FB53, SCL
TITLE = CLK_PULSE
{ S7_Optimized_Access := 'FALSE' }
AUTHOR : hugo
FAMILY : GENERAT
NAME : CLK_PULS